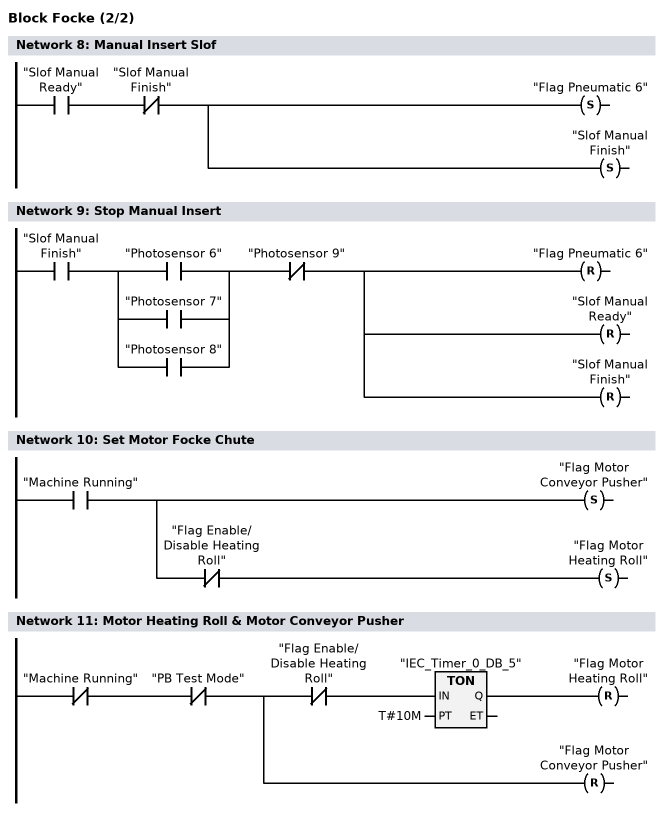
   RUNG wire#powerrail
      Contact( "Slof Manual Ready" )
      I_Contact( "Slof Manual Finish" )
      wire#w1
      S_Coil( "Flag Pneumatic 6" )
   END_RUNG
   RUNG wire#w1
      S_Coil( "Slof Manual Finish" )
   END_RUNG
   // the same network as SCL:
   IF "Slof Manual Ready" AND NOT "Slof Manual Finish" THEN
       "Flag Pneumatic 6" := TRUE;
       "Slof Manual Finish" := TRUE;
   END_IF;
END_REGION

REGION Network 9: Stop Manual Insert
   RUNG wire#powerrail
      Contact( "Slof Manual Finish" )
      wire#w1
      Contact( "Photosensor 6" )
      wire#w2
      I_Contact( "Photosensor 9" )
      wire#w3
      R_Coil( "Flag Pneumatic 6" )
   END_RUNG
   RUNG wire#w1
      Contact( "Photosensor 7" )
   END_RUNG wire#w2
   RUNG wire#w1
      Contact( "Photosensor 8" )
   END_RUNG wire#w2
   RUNG wire#w3
      R_Coil( "Slof Manual Ready" )
   END_RUNG
   RUNG wire#w3
      R_Coil( "Slof Manual Finish" )
   END_RUNG
   // the same network as SCL:
   IF "Slof Manual Finish" AND ("Photosensor 6" OR "Photosensor 7" OR "Photosensor 8") AND NOT "Photosensor 9" THEN
       "Flag Pneumatic 6" := FALSE;
       "Slof Manual Ready" := FALSE;
       "Slof Manual Finish" := FALSE;
   END_IF;
END_REGION

REGION Network 10: Set Motor Focke Chute
   RUNG wire#powerrail
      Contact( "Machine Running" )
      wire#w1
      S_Coil( "Flag Motor Conveyor Pusher" )
   END_RUNG
   RUNG wire#w1
      I_Contact( "Flag Enable/Disable Heating Roll" )
      S_Coil( "Flag Motor Heating Roll" )
   END_RUNG
   // the same network as SCL:
   IF "Machine Running" THEN "Flag Motor Conveyor Pusher" := TRUE; END_IF;
   IF "Machine Running" AND NOT "Flag Enable/Disable Heating Roll" THEN
       "Flag Motor Heating Roll" := TRUE;
   END_IF;
END_REGION

REGION Network 11: Motor Heating Roll & Motor Conveyor Pusher
   #_w1 := NOT "Machine Running" AND NOT "PB Test Mode";
   "IEC_Timer_0_DB_5".TON(IN := #_w1 AND NOT "Flag Enable/Disable Heating Roll", PT := T#10M);
   IF "IEC_Timer_0_DB_5".Q THEN "Flag Motor Heating Roll" := FALSE; END_IF;
   IF #_w1 THEN "Flag Motor Conveyor Pusher" := FALSE; END_IF;
END_REGION
END_FUNCTION_BLOCK

FUNCTION_BLOCK "S Block Par Statistika"   // FB7, LAD
{ S7_Optimized_Access := 'TRUE' }
VERSION : 0.1
BEGIN

REGION Network 1: Move Data Dari HMI Ke Setting Time
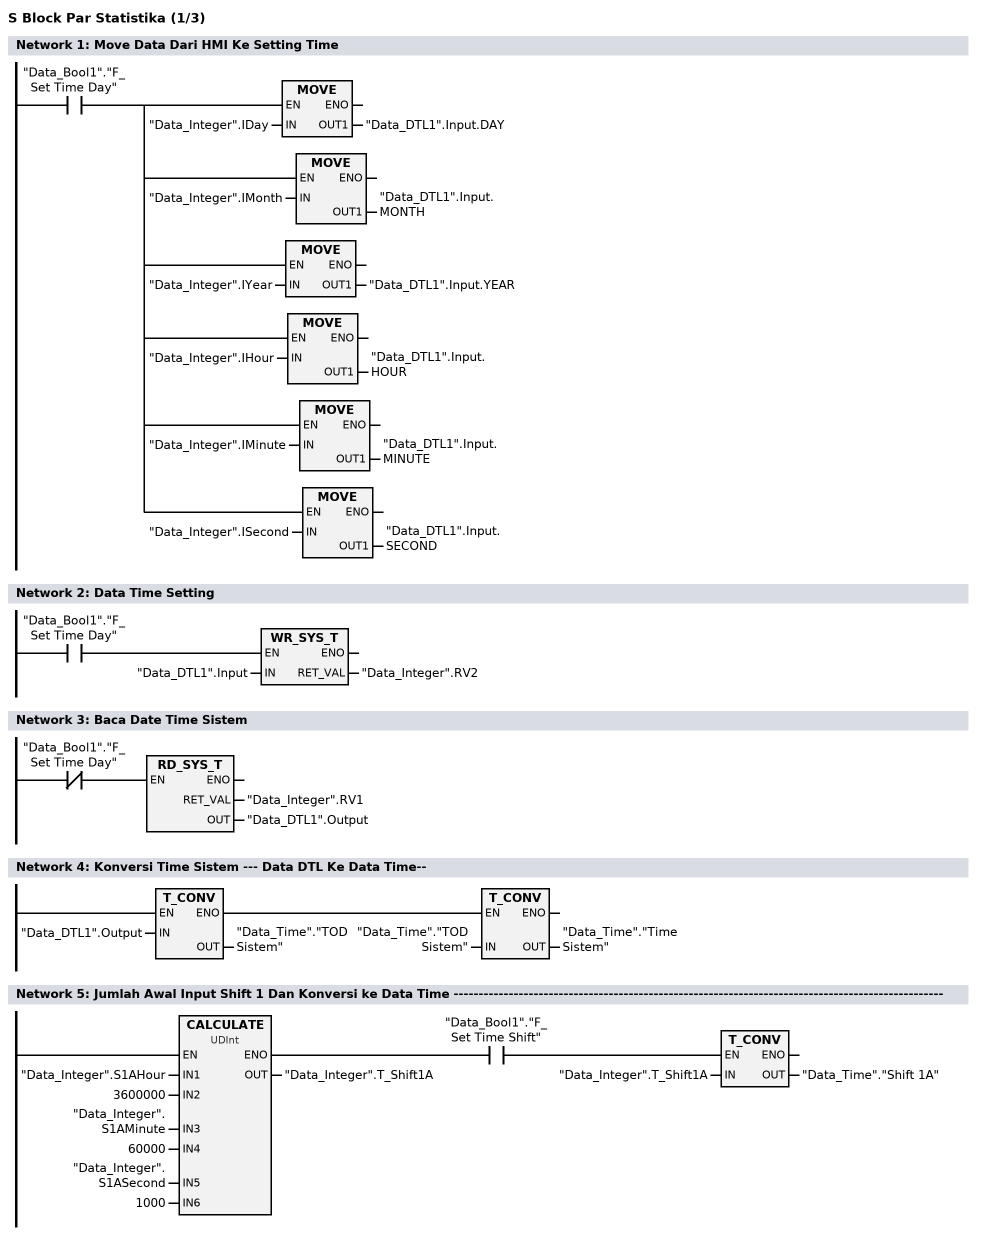
   RUNG wire#powerrail
      Contact( "Data_Bool1"."F_Set Time Day" )
      wire#w1
      { S7_GenerateENO := "TRUE" } Move(in := "Data_Integer".IDay, out1 => "Data_DTL1".Input.DAY)
   END_RUNG
   RUNG wire#w1
      { S7_GenerateENO := "TRUE" } Move(in := "Data_Integer".IMonth, out1 => "Data_DTL1".Input.MONTH)
   END_RUNG
   RUNG wire#w1
      { S7_GenerateENO := "TRUE" } Move(in := "Data_Integer".IYear, out1 => "Data_DTL1".Input.YEAR)
   END_RUNG
   RUNG wire#w1
      { S7_GenerateENO := "TRUE" } Move(in := "Data_Integer".IHour, out1 => "Data_DTL1".Input.HOUR)
   END_RUNG
   RUNG wire#w1
      { S7_GenerateENO := "TRUE" } Move(in := "Data_Integer".IMinute, out1 => "Data_DTL1".Input.MINUTE)
   END_RUNG
   RUNG wire#w1
      { S7_GenerateENO := "TRUE" } Move(in := "Data_Integer".ISecond, out1 => "Data_DTL1".Input.SECOND)
   END_RUNG
   // the same network as SCL:
   IF "Data_Bool1"."F_Set Time Day" THEN
       "Data_DTL1".Input.DAY := "Data_Integer".IDay;
       "Data_DTL1".Input.MONTH := "Data_Integer".IMonth;
       "Data_DTL1".Input.YEAR := "Data_Integer".IYear;
       "Data_DTL1".Input.HOUR := "Data_Integer".IHour;
       "Data_DTL1".Input.MINUTE := "Data_Integer".IMinute;
       "Data_DTL1".Input.SECOND := "Data_Integer".ISecond;
   END_IF;
END_REGION

REGION Network 2: Data Time Setting
   IF "Data_Bool1"."F_Set Time Day" THEN "Data_Integer".RV2 := WR_SYS_T(IN := "Data_DTL1".Input); END_IF;
END_REGION

REGION Network 3: Baca Date Time Sistem
   IF NOT "Data_Bool1"."F_Set Time Day" THEN
       "Data_Integer".RV1 := RD_SYS_T(OUT => "Data_DTL1".Output);
   END_IF;
END_REGION

REGION Network 4: Konversi Time Sistem --- Data DTL Ke Data Time--
   // ENO of a box is taken as its EN; it also drops when the box reports an error
   "Data_Time"."TOD Sistem" := T_CONV(IN := "Data_DTL1".Output);
   "Data_Time"."Time Sistem" := T_CONV(IN := "Data_Time"."TOD Sistem");
END_REGION

REGION Network 5: Jumlah Awal Input Shift 1 Dan Konversi ke Data Time --------------------------------------------------------------------------------------------------
   // ENO of a box is taken as its EN; it also drops when the box reports an error
   "Data_Integer".T_Shift1A := ("Data_Integer".S1AHour*3600000)+("Data_Integer".S1AMinute*60000)+("Data_Integer".S1ASecond*1000);
   IF "Data_Bool1"."F_Set Time Shift" THEN
       "Data_Time"."Shift 1A" := T_CONV(IN := "Data_Integer".T_Shift1A);
   END_IF;
END_REGION

REGION Network 6: Jumlah Akhir Input Shift 1 Dan Konversi ke Data Time @@@@@@@@@@@
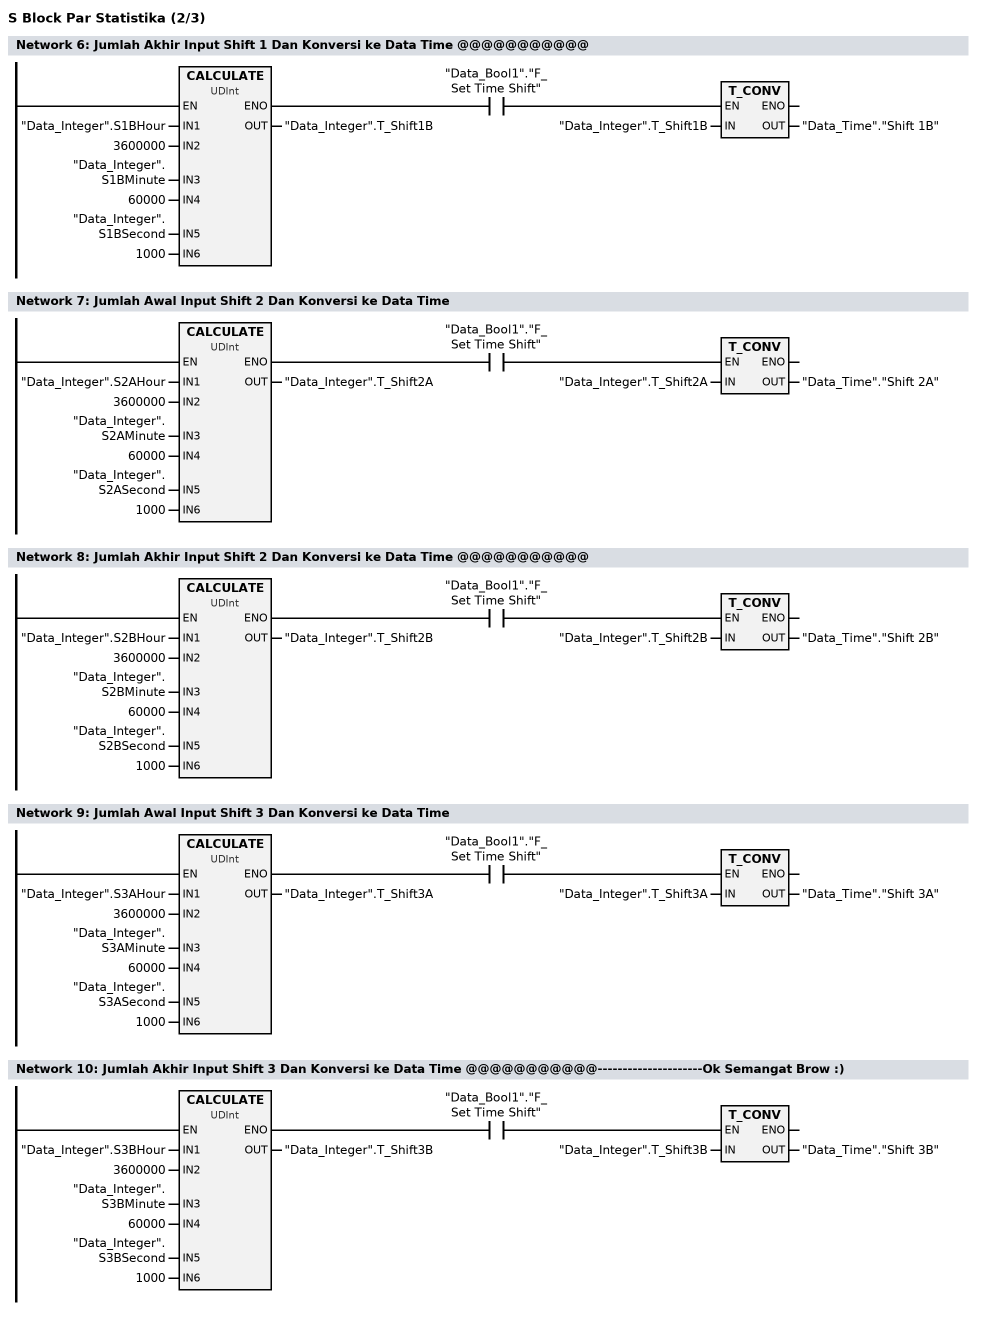
   // ENO of a box is taken as its EN; it also drops when the box reports an error
   "Data_Integer".T_Shift1B := ("Data_Integer".S1BHour*3600000)+("Data_Integer".S1BMinute*60000)+("Data_Integer".S1BSecond*1000);
   IF "Data_Bool1"."F_Set Time Shift" THEN
       "Data_Time"."Shift 1B" := T_CONV(IN := "Data_Integer".T_Shift1B);
   END_IF;
END_REGION

REGION Network 7: Jumlah Awal Input Shift 2 Dan Konversi ke Data Time
   // ENO of a box is taken as its EN; it also drops when the box reports an error
   "Data_Integer".T_Shift2A := ("Data_Integer".S2AHour*3600000)+("Data_Integer".S2AMinute*60000)+("Data_Integer".S2ASecond*1000);
   IF "Data_Bool1"."F_Set Time Shift" THEN
       "Data_Time"."Shift 2A" := T_CONV(IN := "Data_Integer".T_Shift2A);
   END_IF;
END_REGION

REGION Network 8: Jumlah Akhir Input Shift 2 Dan Konversi ke Data Time @@@@@@@@@@@
   // ENO of a box is taken as its EN; it also drops when the box reports an error
   "Data_Integer".T_Shift2B := ("Data_Integer".S2BHour*3600000)+("Data_Integer".S2BMinute*60000)+("Data_Integer".S2BSecond*1000);
   IF "Data_Bool1"."F_Set Time Shift" THEN
       "Data_Time"."Shift 2B" := T_CONV(IN := "Data_Integer".T_Shift2B);
   END_IF;
END_REGION

REGION Network 9: Jumlah Awal Input Shift 3 Dan Konversi ke Data Time
   // ENO of a box is taken as its EN; it also drops when the box reports an error
   "Data_Integer".T_Shift3A := ("Data_Integer".S3AHour*3600000)+("Data_Integer".S3AMinute*60000)+("Data_Integer".S3ASecond*1000);
   IF "Data_Bool1"."F_Set Time Shift" THEN
       "Data_Time"."Shift 3A" := T_CONV(IN := "Data_Integer".T_Shift3A);
   END_IF;
END_REGION

REGION Network 10: Jumlah Akhir Input Shift 3 Dan Konversi ke Data Time @@@@@@@@@@@---------------------Ok Semangat Brow :)
   // ENO of a box is taken as its EN; it also drops when the box reports an error
   "Data_Integer".T_Shift3B := ("Data_Integer".S3BHour*3600000)+("Data_Integer".S3BMinute*60000)+("Data_Integer".S3BSecond*1000);
   IF "Data_Bool1"."F_Set Time Shift" THEN
       "Data_Time"."Shift 3B" := T_CONV(IN := "Data_Integer".T_Shift3B);
   END_IF;
END_REGION

REGION Network 11: Data Time 5 Detik Sebelum Akhir Shift (Waktu Proses Copy Data Current minus 1 sampai 5
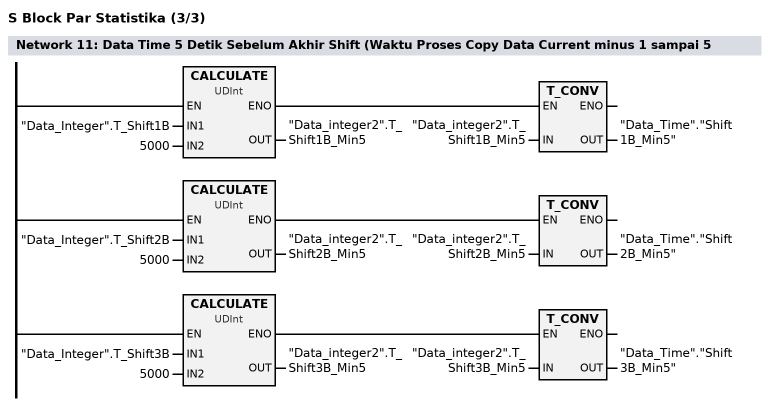
   // ENO of a box is taken as its EN; it also drops when the box reports an error
   "Data_integer2".T_Shift1B_Min5 := "Data_Integer".T_Shift1B-5000;
   "Data_Time"."Shift 1B_Min5" := T_CONV(IN := "Data_integer2".T_Shift1B_Min5);
   "Data_integer2".T_Shift2B_Min5 := "Data_Integer".T_Shift2B-5000;
   "Data_Time"."Shift 2B_Min5" := T_CONV(IN := "Data_integer2".T_Shift2B_Min5);
   "Data_integer2".T_Shift3B_Min5 := "Data_Integer".T_Shift3B-5000;
   "Data_Time"."Shift 3B_Min5" := T_CONV(IN := "Data_integer2".T_Shift3B_Min5);
END_REGION
END_FUNCTION_BLOCK

FUNCTION_BLOCK "S Block Hapus Data"   // FB8, LAD
{ S7_Optimized_Access := 'TRUE' }
VERSION : 0.1
BEGIN

REGION Network 1: Hapus Data Jumlah Sloft Sloft
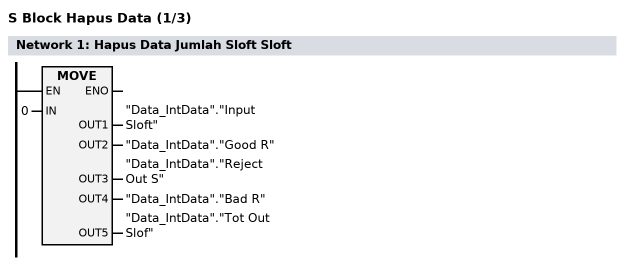
   RUNG wire#powerrail
      { S7_GenerateENO := "TRUE" } Move(in := 0, out1 => "Data_IntData"."Input Sloft", out2 => "Data_IntData"."Good R", out3 => "Data_IntData"."Reject Out S", out4 => "Data_IntData"."Bad R", out5 => "Data_IntData"."Tot Out Slof")
   END_RUNG
   // the same network as SCL:
   "Data_IntData"."Input Sloft" := 0;
   "Data_IntData"."Good R" := 0;
   "Data_IntData"."Reject Out S" := 0;
   "Data_IntData"."Bad R" := 0;
   "Data_IntData"."Tot Out Slof" := 0;
END_REGION

REGION Network 2: Hapus Data Counter Error
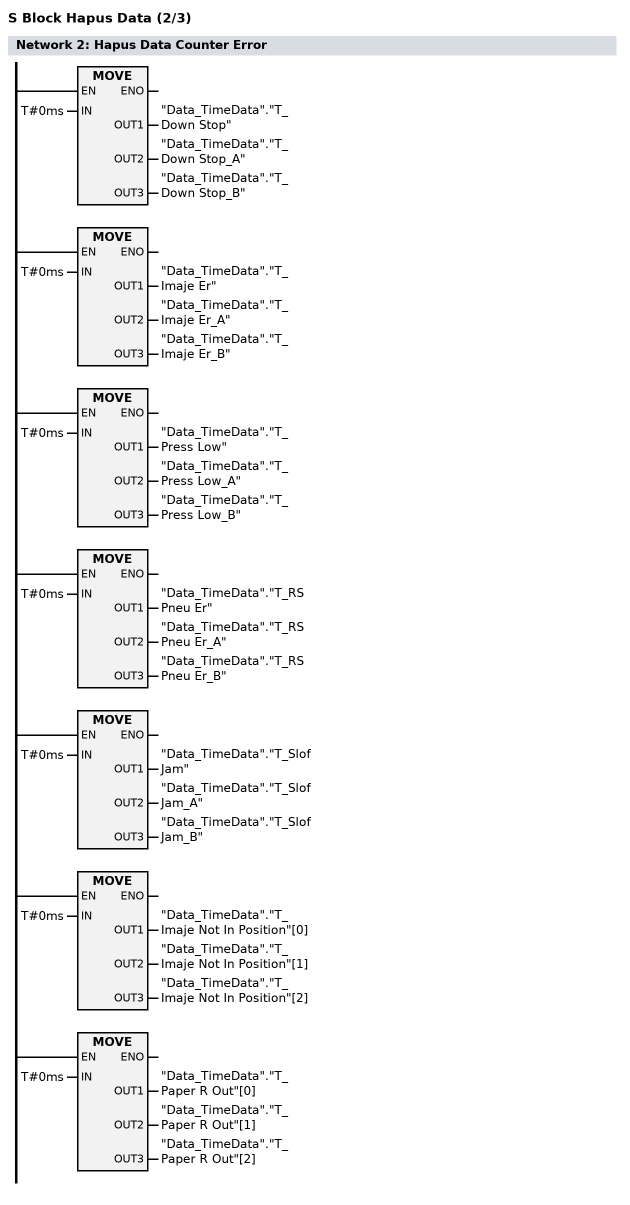
   RUNG wire#powerrail
      { S7_GenerateENO := "TRUE" } Move(in := T#0ms, out1 => "Data_TimeData"."T_Down Stop", out2 => "Data_TimeData"."T_Down Stop_A", out3 => "Data_TimeData"."T_Down Stop_B")
   END_RUNG
   RUNG wire#powerrail
      { S7_GenerateENO := "TRUE" } Move(in := T#0ms, out1 => "Data_TimeData"."T_Imaje Er", out2 => "Data_TimeData"."T_Imaje Er_A", out3 => "Data_TimeData"."T_Imaje Er_B")
   END_RUNG
   RUNG wire#powerrail
      { S7_GenerateENO := "TRUE" } Move(in := T#0ms, out1 => "Data_TimeData"."T_Press Low", out2 => "Data_TimeData"."T_Press Low_A", out3 => "Data_TimeData"."T_Press Low_B")
   END_RUNG
   RUNG wire#powerrail
      { S7_GenerateENO := "TRUE" } Move(in := T#0ms, out1 => "Data_TimeData"."T_RS Pneu Er", out2 => "Data_TimeData"."T_RS Pneu Er_A", out3 => "Data_TimeData"."T_RS Pneu Er_B")
   END_RUNG
   RUNG wire#powerrail
      { S7_GenerateENO := "TRUE" } Move(in := T#0ms, out1 => "Data_TimeData"."T_Slof Jam", out2 => "Data_TimeData"."T_Slof Jam_A", out3 => "Data_TimeData"."T_Slof Jam_B")
   END_RUNG
   RUNG wire#powerrail
      { S7_GenerateENO := "TRUE" } Move(in := T#0ms, out1 => "Data_TimeData"."T_Imaje Not In Position"[0], out2 => "Data_TimeData"."T_Imaje Not In Position"[1], out3 => "Data_TimeData"."T_Imaje Not In Position"[2])
   END_RUNG
   RUNG wire#powerrail
      { S7_GenerateENO := "TRUE" } Move(in := T#0ms, out1 => "Data_TimeData"."T_Paper R Out"[0], out2 => "Data_TimeData"."T_Paper R Out"[1], out3 => "Data_TimeData"."T_Paper R Out"[2])
   END_RUNG
   // the same network as SCL:
   "Data_TimeData"."T_Down Stop" := T#0ms;
   "Data_TimeData"."T_Down Stop_A" := T#0ms;
   "Data_TimeData"."T_Down Stop_B" := T#0ms;
   "Data_TimeData"."T_Imaje Er" := T#0ms;
   "Data_TimeData"."T_Imaje Er_A" := T#0ms;
   "Data_TimeData"."T_Imaje Er_B" := T#0ms;
   "Data_TimeData"."T_Press Low" := T#0ms;
   "Data_TimeData"."T_Press Low_A" := T#0ms;
   "Data_TimeData"."T_Press Low_B" := T#0ms;
   "Data_TimeData"."T_RS Pneu Er" := T#0ms;
   "Data_TimeData"."T_RS Pneu Er_A" := T#0ms;
   "Data_TimeData"."T_RS Pneu Er_B" := T#0ms;
   "Data_TimeData"."T_Slof Jam" := T#0ms;
   "Data_TimeData"."T_Slof Jam_A" := T#0ms;
   "Data_TimeData"."T_Slof Jam_B" := T#0ms;
   "Data_TimeData"."T_Imaje Not In Position"[0] := T#0ms;
   "Data_TimeData"."T_Imaje Not In Position"[1] := T#0ms;
   "Data_TimeData"."T_Imaje Not In Position"[2] := T#0ms;
   "Data_TimeData"."T_Paper R Out"[0] := T#0ms;
   "Data_TimeData"."T_Paper R Out"[1] := T#0ms;
   "Data_TimeData"."T_Paper R Out"[2] := T#0ms;
END_REGION

REGION Network 3: Hapus Data % _____$$$$$$$$$________%
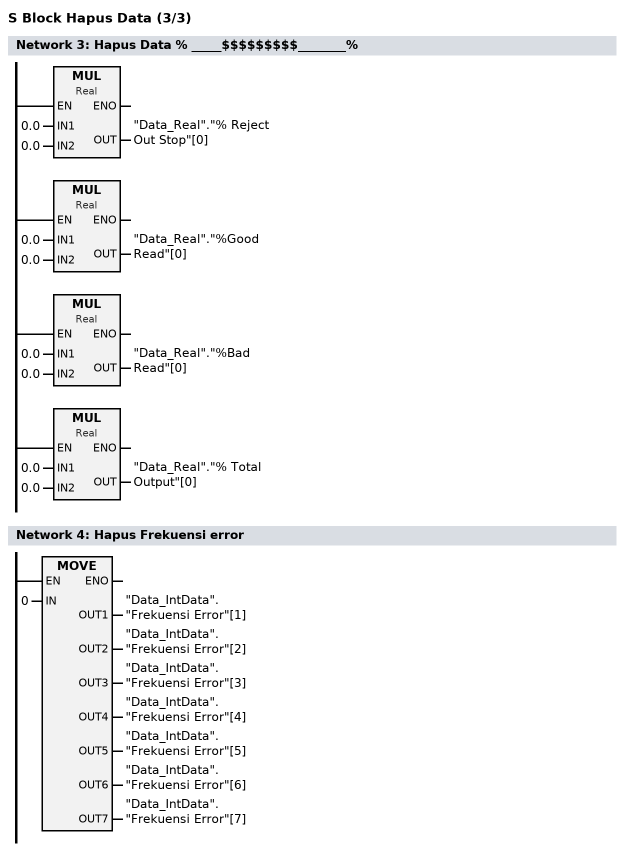
   RUNG wire#powerrail
      { S7_Templates := "SrcType := Real"; S7_GenerateENO := "TRUE" } Mul(in1 := 0.0, in2 := 0.0, out => "Data_Real"."% Reject Out Stop"[0])
   END_RUNG
   RUNG wire#powerrail
      { S7_Templates := "SrcType := Real"; S7_GenerateENO := "TRUE" } Mul(in1 := 0.0, in2 := 0.0, out => "Data_Real"."%Good Read"[0])
   END_RUNG
   RUNG wire#powerrail
      { S7_Templates := "SrcType := Real"; S7_GenerateENO := "TRUE" } Mul(in1 := 0.0, in2 := 0.0, out => "Data_Real"."%Bad Read"[0])
   END_RUNG
   RUNG wire#powerrail
      { S7_Templates := "SrcType := Real"; S7_GenerateENO := "TRUE" } Mul(in1 := 0.0, in2 := 0.0, out => "Data_Real"."% Total Output"[0])
   END_RUNG
   // the same network as SCL:
   "Data_Real"."% Reject Out Stop"[0] := 0.0 * 0.0;
   "Data_Real"."%Good Read"[0] := 0.0 * 0.0;
   "Data_Real"."%Bad Read"[0] := 0.0 * 0.0;
   "Data_Real"."% Total Output"[0] := 0.0 * 0.0;
END_REGION

REGION Network 4: Hapus Frekuensi error
   RUNG wire#powerrail
      { S7_GenerateENO := "TRUE" } Move(in := 0, out1 => "Data_IntData"."Frekuensi Error"[1], out2 => "Data_IntData"."Frekuensi Error"[2], out3 => "Data_IntData"."Frekuensi Error"[3], out4 => "Data_IntData"."Frekuensi Error"[4], out5 => "Data_IntData"."Frekuensi Error"[5], out6 => "Data_IntData"."Frekuensi Error"[6], out7 => "Data_IntData"."Frekuensi Error"[7])
   END_RUNG
   // the same network as SCL:
   "Data_IntData"."Frekuensi Error"[1] := 0;
   "Data_IntData"."Frekuensi Error"[2] := 0;
   "Data_IntData"."Frekuensi Error"[3] := 0;
   "Data_IntData"."Frekuensi Error"[4] := 0;
   "Data_IntData"."Frekuensi Error"[5] := 0;
   "Data_IntData"."Frekuensi Error"[6] := 0;
   "Data_IntData"."Frekuensi Error"[7] := 0;
END_REGION
END_FUNCTION_BLOCK

FUNCTION_BLOCK "S Block Current Shift_M1"   // FB9, LAD
{ S7_Optimized_Access := 'TRUE' }
VERSION : 0.1
BEGIN

REGION Network 1: Move Data Input sloft Minus 0 To 1
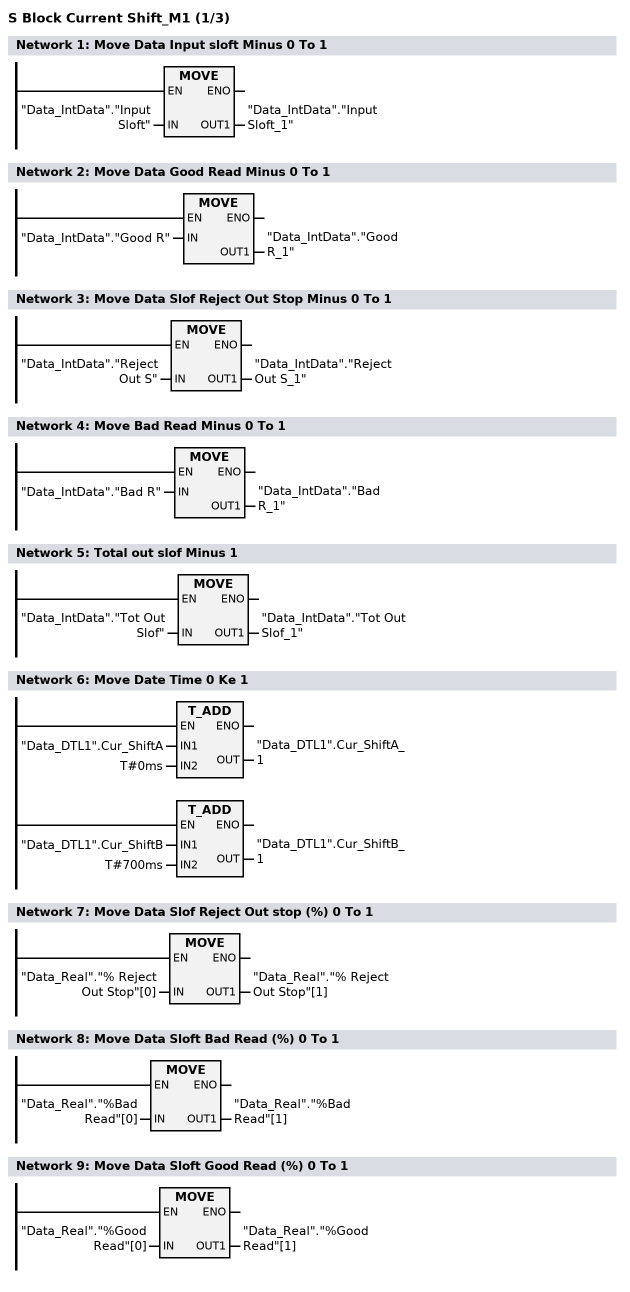
   RUNG wire#powerrail
      { S7_GenerateENO := "TRUE" } Move(in := "Data_IntData"."Input Sloft", out1 => "Data_IntData"."Input Sloft_1")
   END_RUNG
   // the same network as SCL:
   "Data_IntData"."Input Sloft_1" := "Data_IntData"."Input Sloft";
END_REGION

REGION Network 2: Move Data Good Read Minus 0 To 1
   RUNG wire#powerrail
      { S7_GenerateENO := "TRUE" } Move(in := "Data_IntData"."Good R", out1 => "Data_IntData"."Good R_1")
   END_RUNG
   // the same network as SCL:
   "Data_IntData"."Good R_1" := "Data_IntData"."Good R";
END_REGION

REGION Network 3: Move Data Slof Reject Out Stop Minus 0 To 1
   RUNG wire#powerrail
      { S7_GenerateENO := "TRUE" } Move(in := "Data_IntData"."Reject Out S", out1 => "Data_IntData"."Reject Out S_1")
   END_RUNG
   // the same network as SCL:
   "Data_IntData"."Reject Out S_1" := "Data_IntData"."Reject Out S";
END_REGION

REGION Network 4: Move Bad Read Minus 0 To 1
   RUNG wire#powerrail
      { S7_GenerateENO := "TRUE" } Move(in := "Data_IntData"."Bad R", out1 => "Data_IntData"."Bad R_1")
   END_RUNG
   // the same network as SCL:
   "Data_IntData"."Bad R_1" := "Data_IntData"."Bad R";
END_REGION

REGION Network 5: Total out slof Minus 1
   RUNG wire#powerrail
      { S7_GenerateENO := "TRUE" } Move(in := "Data_IntData"."Tot Out Slof", out1 => "Data_IntData"."Tot Out Slof_1")
   END_RUNG
   // the same network as SCL:
   "Data_IntData"."Tot Out Slof_1" := "Data_IntData"."Tot Out Slof";
END_REGION

REGION Network 6: Move Date Time 0 Ke 1
   "Data_DTL1".Cur_ShiftA_1 := T_ADD(IN1 := "Data_DTL1".Cur_ShiftA, IN2 := T#0ms);
   "Data_DTL1".Cur_ShiftB_1 := T_ADD(IN1 := "Data_DTL1".Cur_ShiftB, IN2 := T#700ms);
END_REGION

REGION Network 7: Move Data Slof Reject Out stop (%) 0 To 1
   RUNG wire#powerrail
      { S7_GenerateENO := "TRUE" } Move(in := "Data_Real"."% Reject Out Stop"[0], out1 => "Data_Real"."% Reject Out Stop"[1])
   END_RUNG
   // the same network as SCL:
   "Data_Real"."% Reject Out Stop"[1] := "Data_Real"."% Reject Out Stop"[0];
END_REGION

REGION Network 8: Move Data Sloft Bad Read (%) 0 To 1
   RUNG wire#powerrail
      { S7_GenerateENO := "TRUE" } Move(in := "Data_Real"."%Bad Read"[0], out1 => "Data_Real"."%Bad Read"[1])
   END_RUNG
   // the same network as SCL:
   "Data_Real"."%Bad Read"[1] := "Data_Real"."%Bad Read"[0];
END_REGION

REGION Network 9: Move Data Sloft Good Read (%) 0 To 1
   RUNG wire#powerrail
      { S7_GenerateENO := "TRUE" } Move(in := "Data_Real"."%Good Read"[0], out1 => "Data_Real"."%Good Read"[1])
   END_RUNG
   // the same network as SCL:
   "Data_Real"."%Good Read"[1] := "Data_Real"."%Good Read"[0];
END_REGION

REGION Network 10: Move Output Data Total Sloft (%) 0 To 1
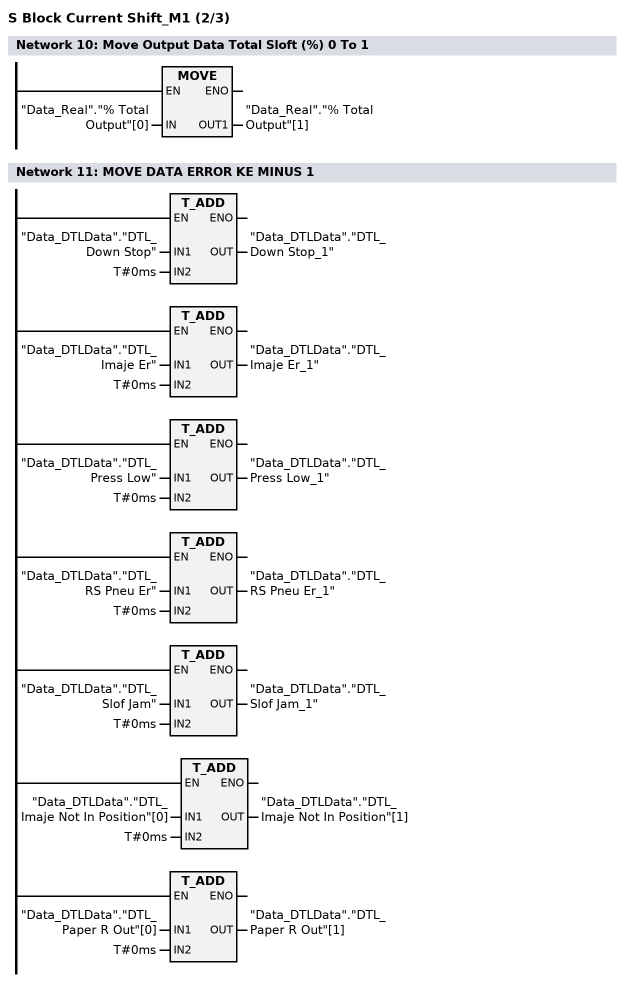
   RUNG wire#powerrail
      { S7_GenerateENO := "TRUE" } Move(in := "Data_Real"."% Total Output"[0], out1 => "Data_Real"."% Total Output"[1])
   END_RUNG
   // the same network as SCL:
   "Data_Real"."% Total Output"[1] := "Data_Real"."% Total Output"[0];
END_REGION

REGION Network 11: MOVE DATA ERROR KE MINUS 1
   "Data_DTLData"."DTL_Down Stop_1" := T_ADD(IN1 := "Data_DTLData"."DTL_Down Stop", IN2 := T#0ms);
   "Data_DTLData"."DTL_Imaje Er_1" := T_ADD(IN1 := "Data_DTLData"."DTL_Imaje Er", IN2 := T#0ms);
   "Data_DTLData"."DTL_Press Low_1" := T_ADD(IN1 := "Data_DTLData"."DTL_Press Low", IN2 := T#0ms);
   "Data_DTLData"."DTL_RS Pneu Er_1" := T_ADD(IN1 := "Data_DTLData"."DTL_RS Pneu Er", IN2 := T#0ms);
   "Data_DTLData"."DTL_Slof Jam_1" := T_ADD(IN1 := "Data_DTLData"."DTL_Slof Jam", IN2 := T#0ms);
   "Data_DTLData"."DTL_Imaje Not In Position"[1] := T_ADD(IN1 := "Data_DTLData"."DTL_Imaje Not In Position"[0],
                           IN2 := T#0ms);
   "Data_DTLData"."DTL_Paper R Out"[1] := T_ADD(IN1 := "Data_DTLData"."DTL_Paper R Out"[0], IN2 := T#0ms);
END_REGION

REGION Network 12: Kopi Jumah Error
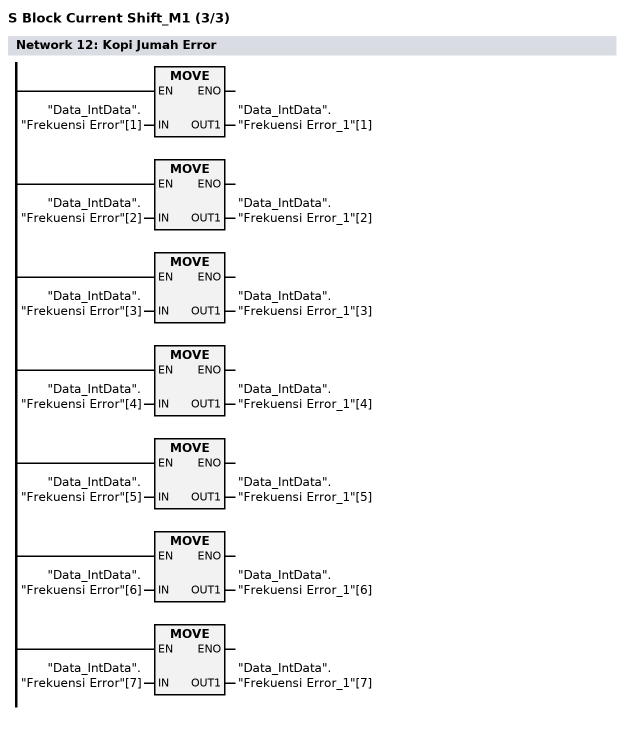
   RUNG wire#powerrail
      { S7_GenerateENO := "TRUE" } Move(in := "Data_IntData"."Frekuensi Error"[1], out1 => "Data_IntData"."Frekuensi Error_1"[1])
   END_RUNG
   RUNG wire#powerrail
      { S7_GenerateENO := "TRUE" } Move(in := "Data_IntData"."Frekuensi Error"[2], out1 => "Data_IntData"."Frekuensi Error_1"[2])
   END_RUNG
   RUNG wire#powerrail
      { S7_GenerateENO := "TRUE" } Move(in := "Data_IntData"."Frekuensi Error"[3], out1 => "Data_IntData"."Frekuensi Error_1"[3])
   END_RUNG
   RUNG wire#powerrail
      { S7_GenerateENO := "TRUE" } Move(in := "Data_IntData"."Frekuensi Error"[4], out1 => "Data_IntData"."Frekuensi Error_1"[4])
   END_RUNG
   RUNG wire#powerrail
      { S7_GenerateENO := "TRUE" } Move(in := "Data_IntData"."Frekuensi Error"[5], out1 => "Data_IntData"."Frekuensi Error_1"[5])
   END_RUNG
   RUNG wire#powerrail
      { S7_GenerateENO := "TRUE" } Move(in := "Data_IntData"."Frekuensi Error"[6], out1 => "Data_IntData"."Frekuensi Error_1"[6])
   END_RUNG
   RUNG wire#powerrail
      { S7_GenerateENO := "TRUE" } Move(in := "Data_IntData"."Frekuensi Error"[7], out1 => "Data_IntData"."Frekuensi Error_1"[7])
   END_RUNG
   // the same network as SCL:
   "Data_IntData"."Frekuensi Error_1"[1] := "Data_IntData"."Frekuensi Error"[1];
   "Data_IntData"."Frekuensi Error_1"[2] := "Data_IntData"."Frekuensi Error"[2];
   "Data_IntData"."Frekuensi Error_1"[3] := "Data_IntData"."Frekuensi Error"[3];
   "Data_IntData"."Frekuensi Error_1"[4] := "Data_IntData"."Frekuensi Error"[4];
   "Data_IntData"."Frekuensi Error_1"[5] := "Data_IntData"."Frekuensi Error"[5];
   "Data_IntData"."Frekuensi Error_1"[6] := "Data_IntData"."Frekuensi Error"[6];
   "Data_IntData"."Frekuensi Error_1"[7] := "Data_IntData"."Frekuensi Error"[7];
END_REGION
END_FUNCTION_BLOCK

FUNCTION_BLOCK "S Check Range Shift"   // FB10, LAD
{ S7_Optimized_Access := 'TRUE' }
VERSION : 0.1
   VAR_TEMP   // added for the SCL form of the ladder/FBD networks
      _w1 : Bool;
      _w2 : Bool;
      _w3 : Bool;
   END_VAR
BEGIN

REGION Network 1: Check Shift 1
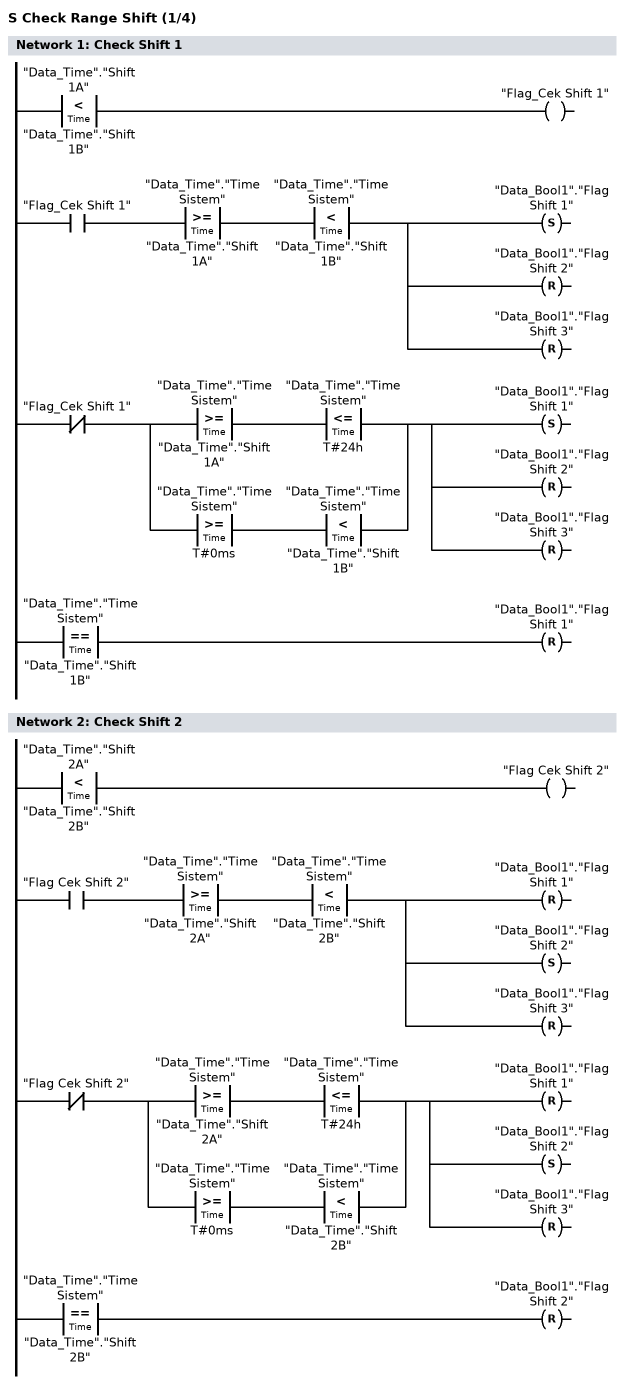
   RUNG wire#powerrail
      { S7_Templates := "SrcType := Time" } LT_Contact(in1 := "Data_Time"."Shift 1A", in2 := "Data_Time"."Shift 1B")
      Coil( "Flag_Cek Shift 1" )
   END_RUNG
   RUNG wire#powerrail
      Contact( "Flag_Cek Shift 1" )
      { S7_Templates := "SrcType := Time" } GE_Contact(in1 := "Data_Time"."Time Sistem", in2 := "Data_Time"."Shift 1A")
      { S7_Templates := "SrcType := Time" } LT_Contact(in1 := "Data_Time"."Time Sistem", in2 := "Data_Time"."Shift 1B")
      wire#w1
      S_Coil( "Data_Bool1"."Flag Shift 1" )
   END_RUNG
   RUNG wire#w1
      R_Coil( "Data_Bool1"."Flag Shift 2" )
   END_RUNG
   RUNG wire#w1
      R_Coil( "Data_Bool1"."Flag Shift 3" )
   END_RUNG
   RUNG wire#powerrail
      I_Contact( "Flag_Cek Shift 1" )
      wire#w2
      { S7_Templates := "SrcType := Time" } GE_Contact(in1 := "Data_Time"."Time Sistem", in2 := "Data_Time"."Shift 1A")
      { S7_Templates := "SrcType := Time" } LE_Contact(in1 := "Data_Time"."Time Sistem", in2 := T#24h)
      wire#w3
      S_Coil( "Data_Bool1"."Flag Shift 1" )
   END_RUNG
   RUNG wire#w2
      { S7_Templates := "SrcType := Time" } GE_Contact(in1 := "Data_Time"."Time Sistem", in2 := T#0ms)
      { S7_Templates := "SrcType := Time" } LT_Contact(in1 := "Data_Time"."Time Sistem", in2 := "Data_Time"."Shift 1B")
   END_RUNG wire#w3
   RUNG wire#w3
      R_Coil( "Data_Bool1"."Flag Shift 2" )
   END_RUNG
   RUNG wire#w3
      R_Coil( "Data_Bool1"."Flag Shift 3" )
   END_RUNG
   RUNG wire#powerrail
      { S7_Templates := "SrcType := Time" } EQ_Contact(in1 := "Data_Time"."Time Sistem", in2 := "Data_Time"."Shift 1B")
      R_Coil( "Data_Bool1"."Flag Shift 1" )
   END_RUNG
   // the same network as SCL:
   "Flag_Cek Shift 1" := "Data_Time"."Shift 1A" < "Data_Time"."Shift 1B";
   IF "Flag_Cek Shift 1" AND ("Data_Time"."Time Sistem" >= "Data_Time"."Shift 1A") AND ("Data_Time"."Time Sistem" < "Data_Time"."Shift 1B") THEN
       "Data_Bool1"."Flag Shift 1" := TRUE;
       "Data_Bool1"."Flag Shift 2" := FALSE;
       "Data_Bool1"."Flag Shift 3" := FALSE;
   END_IF;
   IF NOT "Flag_Cek Shift 1" AND ((("Data_Time"."Time Sistem" >= "Data_Time"."Shift 1A") AND ("Data_Time"."Time Sistem" <= T#24h)) OR (("Data_Time"."Time Sistem" >= T#0ms) AND ("Data_Time"."Time Sistem" < "Data_Time"."Shift 1B"))) THEN
       "Data_Bool1"."Flag Shift 1" := TRUE;
       "Data_Bool1"."Flag Shift 2" := FALSE;
       "Data_Bool1"."Flag Shift 3" := FALSE;
   END_IF;
   IF "Data_Time"."Time Sistem" = "Data_Time"."Shift 1B" THEN "Data_Bool1"."Flag Shift 1" := FALSE; END_IF;
END_REGION

REGION Network 2: Check Shift 2
   RUNG wire#powerrail
      { S7_Templates := "SrcType := Time" } LT_Contact(in1 := "Data_Time"."Shift 2A", in2 := "Data_Time"."Shift 2B")
      Coil( "Flag Cek Shift 2" )
   END_RUNG
   RUNG wire#powerrail
      Contact( "Flag Cek Shift 2" )
      { S7_Templates := "SrcType := Time" } GE_Contact(in1 := "Data_Time"."Time Sistem", in2 := "Data_Time"."Shift 2A")
      { S7_Templates := "SrcType := Time" } LT_Contact(in1 := "Data_Time"."Time Sistem", in2 := "Data_Time"."Shift 2B")
      wire#w1
      R_Coil( "Data_Bool1"."Flag Shift 1" )
   END_RUNG
   RUNG wire#w1
      S_Coil( "Data_Bool1"."Flag Shift 2" )
   END_RUNG
   RUNG wire#w1
      R_Coil( "Data_Bool1"."Flag Shift 3" )
   END_RUNG
   RUNG wire#powerrail
      I_Contact( "Flag Cek Shift 2" )
      wire#w2
      { S7_Templates := "SrcType := Time" } GE_Contact(in1 := "Data_Time"."Time Sistem", in2 := "Data_Time"."Shift 2A")
      { S7_Templates := "SrcType := Time" } LE_Contact(in1 := "Data_Time"."Time Sistem", in2 := T#24h)
      wire#w3
      R_Coil( "Data_Bool1"."Flag Shift 1" )
   END_RUNG
   RUNG wire#w2
      { S7_Templates := "SrcType := Time" } GE_Contact(in1 := "Data_Time"."Time Sistem", in2 := T#0ms)
      { S7_Templates := "SrcType := Time" } LT_Contact(in1 := "Data_Time"."Time Sistem", in2 := "Data_Time"."Shift 2B")
   END_RUNG wire#w3
   RUNG wire#w3
      S_Coil( "Data_Bool1"."Flag Shift 2" )
   END_RUNG
   RUNG wire#w3
      R_Coil( "Data_Bool1"."Flag Shift 3" )
   END_RUNG
   RUNG wire#powerrail
      { S7_Templates := "SrcType := Time" } EQ_Contact(in1 := "Data_Time"."Time Sistem", in2 := "Data_Time"."Shift 2B")
      R_Coil( "Data_Bool1"."Flag Shift 2" )
   END_RUNG
   // the same network as SCL:
   "Flag Cek Shift 2" := "Data_Time"."Shift 2A" < "Data_Time"."Shift 2B";
   IF "Flag Cek Shift 2" AND ("Data_Time"."Time Sistem" >= "Data_Time"."Shift 2A") AND ("Data_Time"."Time Sistem" < "Data_Time"."Shift 2B") THEN
       "Data_Bool1"."Flag Shift 1" := FALSE;
       "Data_Bool1"."Flag Shift 2" := TRUE;
       "Data_Bool1"."Flag Shift 3" := FALSE;
   END_IF;
   IF NOT "Flag Cek Shift 2" AND ((("Data_Time"."Time Sistem" >= "Data_Time"."Shift 2A") AND ("Data_Time"."Time Sistem" <= T#24h)) OR (("Data_Time"."Time Sistem" >= T#0ms) AND ("Data_Time"."Time Sistem" < "Data_Time"."Shift 2B"))) THEN
       "Data_Bool1"."Flag Shift 1" := FALSE;
       "Data_Bool1"."Flag Shift 2" := TRUE;
       "Data_Bool1"."Flag Shift 3" := FALSE;
   END_IF;
   IF "Data_Time"."Time Sistem" = "Data_Time"."Shift 2B" THEN "Data_Bool1"."Flag Shift 2" := FALSE; END_IF;
END_REGION

REGION Network 3: Check Shift 3